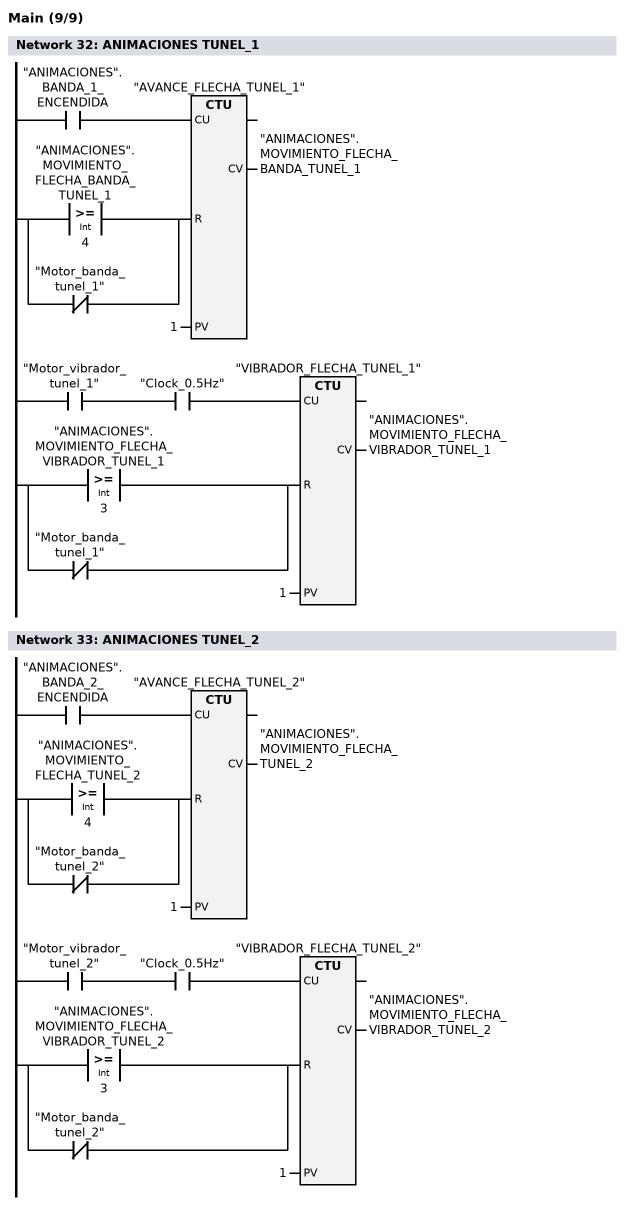
   "AVANCE_FLECHA_TUNEL_1".CTU(CU := "ANIMACIONES".BANDA_1_ENCENDIDA,
                           R := ("ANIMACIONES".MOVIMIENTO_FLECHA_BANDA_TUNEL_1 >= 4) OR NOT "Motor_banda_tunel_1",
                           PV := 1,
                           CV => "ANIMACIONES".MOVIMIENTO_FLECHA_BANDA_TUNEL_1);
   "VIBRADOR_FLECHA_TUNEL_1".CTU(CU := "Motor_vibrador_tunel_1" AND "Clock_0.5Hz",
                           R := ("ANIMACIONES".MOVIMIENTO_FLECHA_VIBRADOR_TUNEL_1 >= 3) OR NOT "Motor_banda_tunel_1",
                           PV := 1,
                           CV => "ANIMACIONES".MOVIMIENTO_FLECHA_VIBRADOR_TUNEL_1);
END_REGION

REGION Network 33: ANIMACIONES TUNEL_2
   "AVANCE_FLECHA_TUNEL_2".CTU(CU := "ANIMACIONES".BANDA_2_ENCENDIDA,
                           R := ("ANIMACIONES".MOVIMIENTO_FLECHA_TUNEL_2 >= 4) OR NOT "Motor_banda_tunel_2",
                           PV := 1,
                           CV => "ANIMACIONES".MOVIMIENTO_FLECHA_TUNEL_2);
   "VIBRADOR_FLECHA_TUNEL_2".CTU(CU := "Motor_vibrador_tunel_2" AND "Clock_0.5Hz",
                           R := ("ANIMACIONES".MOVIMIENTO_FLECHA_VIBRADOR_TUNEL_2 >= 3) OR NOT "Motor_banda_tunel_2",
                           PV := 1,
                           CV => "ANIMACIONES".MOVIMIENTO_FLECHA_VIBRADOR_TUNEL_2);
END_REGION
END_ORGANIZATION_BLOCK

(* ===== HMI "HMI_RT_1" =====
system functions are stored by id; their names below are inferred from use

HMI tags "Default tag table"
   "Tag_ScreenNumber" : UInt, internal

Template "Template_1" 800x480
   Button "Exit" at 714,429 size 71x50; TextOff 'Exit'; PictureOff "ExitRuntime_KTP700_Basic_PN_TR"; PictureOn "ExitRuntime_KTP700_Basic_PN_TR"
      on Release: StopRuntime(0)
   Button "Log on" at 614,429 size 71x50; TextOff 'Log on'; PictureOff "Login_KTP700_Basic_PN_TR"; PictureOn "Login_KTP700_Basic_PN_TR"
      on Release: function_a2a04561()
   Button "Template_Button" at 514,429 size 71x50; TextOff 'Text'
   Button "Template_Button_1" at 414,429 size 71x50; TextOff 'Text'
   Button "Template_Button_2" at 314,429 size 71x50; TextOff 'Text'
   Button "Template_Button_3" at 214,429 size 71x50; TextOff 'Text'
   Button "Alarms" at 114,429 size 71x50; TextOff 'Alarms'; PictureOff "AlarmDisplay_KTP700_Basic_PN_TR"; PictureOn "AlarmDisplay_KTP700_Basic_PN_TR"
      on Release: function_ef3f5d25("Alarm window_Unacknowledged", -1)
   Button "Start screen" at 14,429 size 71x50; TextOff 'Start screen'; PictureOff "NavigateHome_KTP700_Basic_PN_TR"; PictureOn "NavigateHome_KTP700_Basic_PN_TR"
      on Release: ActivateScreen("Root screen", 0)
   SymbolicIOField "Symbolic_IO_Field_Screen" at 93,9 size 600x33; TextOff '0'; TextOn '1'; TextList "TextList_ScreenNames"
      ProcessValue <- "Tag_ScreenNumber"
      on Change: ActivateScreenByNumber("Tag_ScreenNumber", 0)
   DateTimeField "HmiScreenItemData" at 695,25 size 105x25
   DateTimeField "HmiScreenItemData_1" at 695,0 size 105x25
   GraphicView "Logo" at 0,0 size 91x51; Picture "Logo of HMI_1"

screen "Root screen" 800x480, template "Template_1"
   on GenerateScreen: SetTag("Tag_ScreenNumber", 1)
   TextField "HmiScreenItemData" at 80,225 size 640x25; Text 'Welcome to HMI_1 (KTP700 Basic+ PN)!'
*)

(* ===== HMI "HMI_RT_2" =====
system functions are stored by id; their names below are inferred from use
connection "HMI_Connection_1": ETHERNET, SMART_S7_1500_OMS

HMI tags "Default tag table"
   "Tag_ScreenNumber" : UInt, internal
   "Motor_banda_tunel_1" : Bool = PLC Motor_banda_tunel_1 AT %Q10.0, 1 s
   "Señal_de_fallo_banda_tunel_1" : Bool = PLC Señal_de_fallo_banda_tunel_1 AT %I11.1, 1 s
   "PERMISOS_DE_MARCHA_TUNEL_1_BANDA_TUNEL_1_MANUAL" : Bool = PLC PERMISOS_DE_MARCHA_TUNEL_1.BANDA_TUNEL_1_MANUAL, 1 s
   "BOTONERA_HMI_TUNEL_1_KM1_INICIO_MANUAL_BANDA_TUNEL_1" : Bool = PLC BOTONERA_HMI_TUNEL_1.KM1_INICIO_MANUAL_BANDA_TUNEL_1, 1 s
   "BOTONERA_HMI_TUNEL_1_KM1_STOP_MANUAL_BANDA_TUNEL_1" : Bool = PLC BOTONERA_HMI_TUNEL_1.KM1_STOP_MANUAL_BANDA_TUNEL_1, 1 s
   "PERMISOS_DE_MARCHA_TUNEL_1_VENTILADOR_TUNEL_1_MANUAL" : Bool = PLC PERMISOS_DE_MARCHA_TUNEL_1.VENTILADOR_TUNEL_1_MANUAL, 1 s
   "Señal_de_fallo_ventilador_tunel_1" : Bool = PLC Señal_de_fallo_ventilador_tunel_1 AT %I11.3, 1 s
   "BOTONERA_HMI_TUNEL_1_KM2_INICIO_MANUAL_ASPIRADOR_TUNEL_1" : Bool = PLC BOTONERA_HMI_TUNEL_1.KM2_INICIO_MANUAL_ASPIRADOR_TUNEL_1, 1 s
   "BOTONERA_HMI_TUNEL_1_KM3_INICIO_MANUAL_VENTILADOR_TUNEL_1" : Bool = PLC BOTONERA_HMI_TUNEL_1.KM3_INICIO_MANUAL_VENTILADOR_TUNEL_1, 1 s
   "BOTONERA_HMI_TUNEL_1_KM3_STOP_MANUAL_VENTILADOR_TUNEL_1" : Bool = PLC BOTONERA_HMI_TUNEL_1.KM3_STOP_MANUAL_VENTILADOR_TUNEL_1, 1 s
   "PERMISOS_DE_MARCHA_TUNEL_1_ASPIRADOR_TUNEL_1_MANUAL" : Bool = PLC PERMISOS_DE_MARCHA_TUNEL_1.ASPIRADOR_TUNEL_1_MANUAL, 1 s
   "Señal_de_fallo_aspirador_tunel_1" : Bool = PLC Señal_de_fallo_aspirador_tunel_1 AT %I11.2, 1 s
   "BOTONERA_HMI_TUNEL_1_KM2_STOP_MANUAL_ASPIRADOR_TUNEL_1" : Bool = PLC BOTONERA_HMI_TUNEL_1.KM2_STOP_MANUAL_ASPIRADOR_TUNEL_1, 1 s
   "PERMISOS_DE_MARCHA_TUNEL_1_CERRAR_CUCHARA_TUNEL_1_MANUAL" : Bool = PLC PERMISOS_DE_MARCHA_TUNEL_1.CERRAR_CUCHARA_TUNEL_1_MANUAL, 1 s
   "PERMISOS_DE_MARCHA_TUNEL_1_ABRIR_CUCHARA_TUNEL_1_MANUAL" : Bool = PLC PERMISOS_DE_MARCHA_TUNEL_1.ABRIR_CUCHARA_TUNEL_1_MANUAL, 1 s
   "BOTONERA_HMI_TUNEL_1_SUBIR_CUCHARA_TUNEL_1" : Bool = PLC BOTONERA_HMI_TUNEL_1.SUBIR_CUCHARA_TUNEL_1, 1 s
   "BOTONERA_HMI_TUNEL_1_BAJAR_CUCHARA_TUNEL_1" : Bool = PLC BOTONERA_HMI_TUNEL_1.BAJAR_CUCHARA_TUNEL_1, 1 s
   "BOTONERA_HMI_TUNEL_1_CARGADOR_CAJAS_IZQUIERDA_TUNEL_1" : Bool = PLC BOTONERA_HMI_TUNEL_1.CARGADOR_CAJAS_IZQUIERDA_TUNEL_1, 1 s
   "PERMISOS_DE_MARCHA_TUNEL_1_CAJA_IZQUIERDA_TUNEL_1_MANUAL" : Bool = PLC PERMISOS_DE_MARCHA_TUNEL_1.CAJA_IZQUIERDA_TUNEL_1_MANUAL, 1 s
   "PERMISOS_DE_MARCHA_TUNEL_1_CAJA_DERECHA_TUNEL_1_MANUAL" : Bool = PLC PERMISOS_DE_MARCHA_TUNEL_1.CAJA_DERECHA_TUNEL_1_MANUAL, 1 s
   "BOTONERA_HMI_TUNEL_1_CARGADOR_CAJAS_DERECHA_TUNEL_1" : Bool = PLC BOTONERA_HMI_TUNEL_1.CARGADOR_CAJAS_DERECHA_TUNEL_1, 1 s
   "BOTONERA_HMI_TUNEL_1_KM4_INICIO_MANUAL_VIBRADOR_TUNEL_1" : Bool = PLC BOTONERA_HMI_TUNEL_1.KM4_INICIO_MANUAL_VIBRADOR_TUNEL_1, 1 s
   "BOTONERA_HMI_TUNEL_1_KM4_STOP_MANUAL_VIBRADOR_TUNEL_1" : Bool = PLC BOTONERA_HMI_TUNEL_1.KM4_STOP_MANUAL_VIBRADOR_TUNEL_1, 1 s
   "PERMISOS_DE_MARCHA_TUNEL_1_VIBRADOR_TUNEL_1_MANUAL" : Bool = PLC PERMISOS_DE_MARCHA_TUNEL_1.VIBRADOR_TUNEL_1_MANUAL, 1 s
   "Señal_de_fallo_vibrador_tunel_1" : Bool = PLC Señal_de_fallo_vibrador_tunel_1 AT %I11.4, 1 s
   "ANIMACIONES_MOVIMIENTO_FLECHA_TUNEL_1" : Int = PLC ANIMACIONES.MOVIMIENTO_FLECHA_BANDA_TUNEL_1, 1 s
   "ANIMACIONES_MOVIMIENTO_FLECHA_VIBRADOR_TUNEL_1" : Int = PLC ANIMACIONES.MOVIMIENTO_FLECHA_VIBRADOR_TUNEL_1, 1 s
   "Señalizacion_operacion_verde_tunel_1" : Bool = PLC Señalizacion_operacion_verde_tunel_1 AT %Q11.3, 1 s
   "Señalizacion_azul_tunel_1" : Bool = PLC Señalizacion_azul_tunel_1 AT %Q11.2, 1 s
   "Señalizacion_Roja_Tunel_1" : Bool = PLC Señalizacion_Roja_Tunel_1 AT %Q11.1, 1 s
   "PERMISOS_DE_MARCHA_TUNEL_1_VENTILADOR_TUNEL_1_AUTOMATICO" : Bool = PLC PERMISOS_DE_MARCHA_TUNEL_1.VENTILADOR_TUNEL_1_AUTOMATICO, 1 s
   "PERMISOS_DE_MARCHA_TUNEL_1_ASPIRADOR_TUNEL_1_AUTOMATICO" : Bool = PLC PERMISOS_DE_MARCHA_TUNEL_1.ASPIRADOR_TUNEL_1_AUTOMATICO, 1 s
   "PERMISOS_DE_MARCHA_TUNEL_1_BANDA_TUNEL_1_AUTOMATICO" : Bool = PLC PERMISOS_DE_MARCHA_TUNEL_1.BANDA_TUNEL_1_AUTOMATICO, 1 s
   "PERMISOS_DE_MARCHA_TUNEL_1_VIBRADOR_TUNEL_1_AUTOMATICO" : Bool = PLC PERMISOS_DE_MARCHA_TUNEL_1.VIBRADOR_TUNEL_1_AUTOMATICO, 1 s
   "PERMISOS_DE_MARCHA_TUNEL_1_CAJA_DERECHA_TUNEL_1_AUTOMATICO" : Bool = PLC PERMISOS_DE_MARCHA_TUNEL_1.CAJA_DERECHA_TUNEL_1_AUTOMATICO, 1 s
   "PERMISOS_DE_MARCHA_TUNEL_1_CAJA_IZQUIERDA_TUNEL_1_AUTOMATICO" : Bool = PLC PERMISOS_DE_MARCHA_TUNEL_1.CAJA_IZQUIERDA_TUNEL_1_AUTOMATICO, 1 s
   "PERMISOS_DE_MARCHA_TUNEL_1_CERRAR_CUCHARA_TUNEL_1_AUTOMATICO" : Bool = PLC PERMISOS_DE_MARCHA_TUNEL_1.CERRAR_CUCHARA_TUNEL_1_AUTOMATICO, 1 s
   "PERMISOS_DE_MARCHA_TUNEL_1_ABRIR_CUCHARA_TUNEL_1_AUTOMATICO" : Bool = PLC PERMISOS_DE_MARCHA_TUNEL_1.ABRIR_CUCHARA_TUNEL_1_AUTOMATICO, 1 s
   "Motor_aspirador_tunel_!" : Bool = PLC Motor_aspirador_tunel_! AT %Q10.1, 1 s
   "Motor_ventilador_tunel_1" : Bool = PLC Motor_ventilador_tunel_1 AT %Q10.2, 1 s
   "Motor_vibrador_tunel_1" : Bool = PLC Motor_vibrador_tunel_1 AT %Q10.3, 1 s
   "Subir_Cuchara_Tunel_1" : Bool = PLC Subir_Cuchara_Tunel_1 AT %Q11.0, 1 s
   "Bajar_cuchara_Tunel_1" : Bool = PLC Bajar_cuchara_Tunel_1 AT %Q10.7, 1 s
   "Desviar_cajas_derecha_Tunel_1" : Bool = PLC Desviar_cajas_derecha_Tunel_1 AT %Q10.4, 1 s
   "Desviar_cajas_izquierda_Tunel_1" : Bool = PLC Desviar_cajas_izquierda_Tunel_1 AT %Q10.5, 1 s
   "TEMPORIZADOR_PASO_TAPAS_TUNEL_1" : Int = PLC TEMPORIZADOR_PASO_TAPAS_TUNEL_1 AT %MW0, 1 s
   "TEMPORIZADOR_BLOQUEO_TAPAS_TUNEL_1" : Int = PLC TEMPORIZADOR_BLOQUEO_TAPAS_TUNEL_1 AT %MW2, 1 s
   "TEMPORIZADOR_CAMBIO_DE_LLENADO_CAJA_TUNEL_1" : Int = PLC TEMPORIZADOR_CAMBIO_DE_LLENADO_CAJA_TUNEL_1 AT %MW4, 1 s
   "PERMISOS_GENERALES_MODO_LOCAL_1" : Bool = PLC PERMISOS_GENERALES.MODO_LOCAL_1, 1 s
   "PERMISOS_GENERALES_MODO_AUTOMATICO_1" : Bool = PLC PERMISOS_GENERALES.MODO_AUTOMATICO_1, 1 s
   "ALARMAS_TUNEL_1" : Int AT %DB24.DBW0, 1 s

discrete alarms
   1: 'Revisar estado guardamotor QM1', class Errors, trigger "ALARMAS_TUNEL_1" bit 8
   2: 'Revisar estado guardamotor QM2', class Warnings, trigger "ALARMAS_TUNEL_1" bit 9
   3: 'Revisar estado guardamotor QM3', class Warnings, trigger "ALARMAS_TUNEL_1" bit 10
   4: 'Revisar estado guardamotor QM4', class Errors, trigger "ALARMAS_TUNEL_1" bit 11
   5: 'Revisar presion en red neumatica', class Errors, trigger "ALARMAS_TUNEL_1" bit 12
   6: 'Equipo en paro de emergencia', class Errors, trigger "ALARMAS_TUNEL_1" bit 14
   7: 'Sin suministro de tapas en entrada', class Warnings, trigger "ALARMAS_TUNEL_1" bit 13

Template "Template_1" 800x480
   Button "Exit" at 714,429 size 71x50; TextOff 'Exit'; PictureOff "ExitRuntime_KTP700_Basic_PN_TR"; PictureOn "ExitRuntime_KTP700_Basic_PN_TR"
      on Release: StopRuntime(0)
   Button "Log on" at 614,429 size 71x50; TextOff 'Log on'; PictureOff "Login_KTP700_Basic_PN_TR"; PictureOn "Login_KTP700_Basic_PN_TR"
      on Release: function_a2a04561()
   Button "Template_Button" at 514,429 size 71x50; TextOff 'Text'
   Button "Template_Button_1" at 414,429 size 71x50; TextOff 'Text'
   Button "Template_Button_2" at 314,429 size 71x50; TextOff 'Text'
   Button "Template_Button_3" at 214,429 size 71x50; TextOff 'Text'
   Button "Alarms" at 114,429 size 71x50; TextOff 'Alarms'; PictureOff "AlarmDisplay_KTP700_Basic_PN_TR"; PictureOn "AlarmDisplay_KTP700_Basic_PN_TR"
   Button "Start screen" at 14,429 size 71x50; TextOff 'Start screen'; PictureOff "NavigateHome_KTP700_Basic_PN_TR"; PictureOn "NavigateHome_KTP700_Basic_PN_TR"
      on Release: ActivateScreen("PANTALLA DE INICIO", 0)
   SymbolicIOField "Symbolic_IO_Field_Screen" at 93,9 size 600x33; TextOff '0'; TextOn '1'; TextList "TextList_ScreenNames"
      ProcessValue <- "Tag_ScreenNumber"
      on Change: ActivateScreenByNumber("Tag_ScreenNumber", 0)
   DateTimeField "HmiScreenItemData" at 695,25 size 105x25
   DateTimeField "HmiScreenItemData_1" at 695,0 size 105x25
   GraphicView "Logo" at 0,0 size 91x51; Picture "Logo of HMI_1"

screen "PANTALLA DE INICIO" 800x480, template "Template_1"
   on GenerateScreen: SetTag("Tag_ScreenNumber", 1)
   GraphicView "Graphic view_1" at 302,101 size 200x200; Picture "pngegg"
   Button "Button_1" at 277,47 size 251x30; TextOff 'TUNEL ENFRIAMIENTO 1'
   Button "Button_2" at 244,83 size 316x30; TextOff 'LINEA DE FABRICACION DE TAPAS 2'
   GraphicView "Graphic view_2" at 352,314 size 100x100; Picture "selector-de-llave-3-posiciones-enclavamiento-eaton-moeller-111774-m22-wrs3-ms3-removebg-preview"
   Button "Button_3" at 131,282 size 96x32; TextOff 'LOCAL'; Authorization "Mantenimiento"
      on Press: ActivateScreen("MODO LOCAL", 0)
   Button "Button_4" at 590,282 size 96x32; TextOff 'REMOTO'
      on Press: ActivateScreen("MODO REMOTO", 0)

screen "MODO LOCAL" 800x480
   GraphicView "Graphic view_8" at 402,218 size 50x50; Picture "Graphic_9"
      Visibility <- "PERMISOS_DE_MARCHA_TUNEL_1_VENTILADOR_TUNEL_1_MANUAL"
   GraphicView "Graphic view_1" at 0,0 size 100x100; Picture "pngegg"
   GraphicView "Graphic view_2" at 126,262 size 624x99; Picture "Graphic_1"
   GraphicView "Graphic view_3" at 470,311 size 50x50; Picture "Graphic_2"
      Visibility <- "PERMISOS_DE_MARCHA_TUNEL_1_BANDA_TUNEL_1_MANUAL"
   GraphicView "Graphic view_4" at 470,311 size 50x50; Picture "Graphic_3"
      Visibility <- "Motor_banda_tunel_1"
   GraphicView "Graphic view_5" at 470,311 size 50x50; Picture "Graphic_4"
      Visibility <- "Señal_de_fallo_banda_tunel_1"
   Button "Button_2" at 466,363 size 50x20; TextOff 'ON'; Authorization "Mantenimiento"
      on Press: SetBit("BOTONERA_HMI_TUNEL_1_KM1_INICIO_MANUAL_BANDA_TUNEL_1")
      on Release: ResetBit("BOTONERA_HMI_TUNEL_1_KM1_INICIO_MANUAL_BANDA_TUNEL_1")
      Visibility <- "PERMISOS_GENERALES_MODO_LOCAL_1"
   Button "Button_3" at 522,362 size 50x20; TextOff 'OFF'; Authorization "Mantenimiento"
      on Press: SetBit("BOTONERA_HMI_TUNEL_1_KM1_STOP_MANUAL_BANDA_TUNEL_1")
      on Release: ResetBit("BOTONERA_HMI_TUNEL_1_KM1_STOP_MANUAL_BANDA_TUNEL_1")
      Visibility <- "PERMISOS_GENERALES_MODO_LOCAL_1"
   GraphicView "Graphic view_6" at 401,217 size 50x50; Picture "Graphic_6"
      Visibility <- "PERMISOS_DE_MARCHA_TUNEL_1_VENTILADOR_TUNEL_1_MANUAL"
   GraphicView "Graphic view_9" at 356,222 size 48x45; Picture "viento"
      Visibility <- "PERMISOS_DE_MARCHA_TUNEL_1_VENTILADOR_TUNEL_1_MANUAL"
   GraphicView "Graphic view_7" at 401,218 size 50x50; Picture "Graphic_7"
      Visibility <- "Señal_de_fallo_ventilador_tunel_1"
   Button "Button_1" at 359,194 size 50x20; TextOff 'ON'; Authorization "Mantenimiento"
      on Release: ResetBit("BOTONERA_HMI_TUNEL_1_KM3_INICIO_MANUAL_VENTILADOR_TUNEL_1")
      on Press: SetBit("BOTONERA_HMI_TUNEL_1_KM3_INICIO_MANUAL_VENTILADOR_TUNEL_1")
   Button "Button_4" at 419,195 size 50x20; TextOff 'OFF'; Authorization "Mantenimiento"
      on Release: ResetBit("BOTONERA_HMI_TUNEL_1_KM3_STOP_MANUAL_VENTILADOR_TUNEL_1")
      on Press: SetBit("BOTONERA_HMI_TUNEL_1_KM3_STOP_MANUAL_VENTILADOR_TUNEL_1")
   GraphicView "Graphic view_10" at 240,300 size 50x50; Picture "Graphic_23"
      Visibility <- "PERMISOS_DE_MARCHA_TUNEL_1_ASPIRADOR_TUNEL_1_MANUAL"
   GraphicView "Graphic view_11" at 240,300 size 50x50; Picture "Graphic_24"
      Visibility <- "PERMISOS_DE_MARCHA_TUNEL_1_ASPIRADOR_TUNEL_1_MANUAL"
   GraphicView "Graphic view_12" at 240,300 size 50x50; Picture "Graphic_25"
      Visibility <- "Señal_de_fallo_aspirador_tunel_1"
   GraphicView "Graphic view_13" at 209,321 size 52x87; Picture "viento"
      Visibility <- "PERMISOS_DE_MARCHA_TUNEL_1_ASPIRADOR_TUNEL_1_MANUAL"
   Button "Button_5" at 211,388 size 50x20; TextOff 'ON'; Authorization "Mantenimiento"
      on Release: ResetBit("BOTONERA_HMI_TUNEL_1_KM2_INICIO_MANUAL_ASPIRADOR_TUNEL_1")
      on Press: SetBit("BOTONERA_HMI_TUNEL_1_KM2_INICIO_MANUAL_ASPIRADOR_TUNEL_1")
   Button "Button_6" at 265,389 size 50x20; TextOff 'OFF'; Authorization "Mantenimiento"
      on Release: ResetBit("BOTONERA_HMI_TUNEL_1_KM2_STOP_MANUAL_ASPIRADOR_TUNEL_1")
      on Press: SetBit("BOTONERA_HMI_TUNEL_1_KM2_STOP_MANUAL_ASPIRADOR_TUNEL_1")
   TextField "Text field_1" at 463,386 size 109x23; Text 'Motor Banda'
   TextField "Text field_2" at 376,159 size 90x23; Text 'Ventilador'
   TextField "Text field_3" at 231,411 size 81x23; Text 'Extractor'
   GraphicView "Graphic view_15" at 500,76 size 300x200; Picture "Compuerta"
      Visibility <- "PERMISOS_DE_MARCHA_TUNEL_1_ABRIR_CUCHARA_TUNEL_1_MANUAL"
   GraphicView "Graphic view_14" at 499,139 size 300x200; Picture "Compuerta"
      Visibility <- "PERMISOS_DE_MARCHA_TUNEL_1_CERRAR_CUCHARA_TUNEL_1_MANUAL"
   Button "Button_7" at 724,120 size 60x20; TextOff 'SUBIR'; Authorization "Mantenimiento"
      on Release: ResetBit("BOTONERA_HMI_TUNEL_1_SUBIR_CUCHARA_TUNEL_1")
      on Press: SetBit("BOTONERA_HMI_TUNEL_1_SUBIR_CUCHARA_TUNEL_1")
      Appearance <- "PERMISOS_DE_MARCHA_TUNEL_1_ABRIR_CUCHARA_TUNEL_1_MANUAL"
   Button "Button_8" at 724,154 size 60x20; TextOff 'BAJAR'; Authorization "Mantenimiento"
      on Release: ResetBit("BOTONERA_HMI_TUNEL_1_BAJAR_CUCHARA_TUNEL_1")
      on Press: SetBit("BOTONERA_HMI_TUNEL_1_BAJAR_CUCHARA_TUNEL_1")
      Appearance <- "PERMISOS_DE_MARCHA_TUNEL_1_CERRAR_CUCHARA_TUNEL_1_MANUAL"
   Button "Button_9" at 16,155 size 100x20; TextOff 'IZQUIERDA'; Authorization "Mantenimiento"
      on Release: ResetBit("BOTONERA_HMI_TUNEL_1_CARGADOR_CAJAS_IZQUIERDA_TUNEL_1")
      on Press: SetBit("BOTONERA_HMI_TUNEL_1_CARGADOR_CAJAS_IZQUIERDA_TUNEL_1")
      Appearance <- "PERMISOS_DE_MARCHA_TUNEL_1_CAJA_IZQUIERDA_TUNEL_1_MANUAL"
   Button "Button_10" at 169,155 size 100x20; TextOff 'DERECHA'; Authorization "Mantenimiento"
      on Release: ResetBit("BOTONERA_HMI_TUNEL_1_CARGADOR_CAJAS_DERECHA_TUNEL_1")
      on Press: SetBit("BOTONERA_HMI_TUNEL_1_CARGADOR_CAJAS_DERECHA_TUNEL_1")
      Appearance <- "PERMISOS_DE_MARCHA_TUNEL_1_CAJA_DERECHA_TUNEL_1_MANUAL"
   Button "Button_11" at 400,440 size 368x32; TextOff 'ESTADO DE ELEMENTOS Y ACTUADORES'
      on Press: ActivateScreen("VISUALIZACION DE ESTADOS LOCAL TUNEL 1", 0)
   TextField "Text field_4" at 229,86 size 241x33; Text 'MODO LOCAL ACTIVO'
   GraphicView "Graphic view_16" at 496,268 size 87x56; Picture "pngtree-vector-back-icon-png-image_956547-removebg-preview"
      Visibility <- "ANIMACIONES_MOVIMIENTO_FLECHA_TUNEL_1"
   GraphicView "Graphic view_17" at 210,262 size 87x56; Picture "pngtree-vector-back-icon-png-image_956547-removebg-preview"
      Visibility <- "ANIMACIONES_MOVIMIENTO_FLECHA_TUNEL_1"
   GraphicView "Graphic view_18" at 350,266 size 87x56; Picture "pngtree-vector-back-icon-png-image_956547-removebg-preview"
      Visibility <- "ANIMACIONES_MOVIMIENTO_FLECHA_TUNEL_1"
   GraphicView "Graphic view_19" at 0,296 size 209x184; Picture "AGITADOR"
   GraphicView "Graphic view_20" at 16,418 size 50x50; Picture "Graphic_4"
      Visibility <- "Señal_de_fallo_vibrador_tunel_1"
   GraphicView "Graphic view_21" at 16,417 size 50x50; Picture "Graphic_2"
      Visibility <- "PERMISOS_DE_MARCHA_TUNEL_1_VIBRADOR_TUNEL_1_MANUAL"
   GraphicView "Graphic view_22" at 16,416 size 50x50; Picture "Graphic_3"
      Visibility <- "PERMISOS_DE_MARCHA_TUNEL_1_VIBRADOR_TUNEL_1_MANUAL"
   GraphicView "Graphic view_23" at 4,366 size 35x40; Picture "FLECHA ARRIBA"
      Visibility <- "ANIMACIONES_MOVIMIENTO_FLECHA_VIBRADOR_TUNEL_1"
   GraphicView "Graphic view_24" at 160,366 size 35x40; Picture "FLECHA ABAJO"
      Visibility <- "ANIMACIONES_MOVIMIENTO_FLECHA_VIBRADOR_TUNEL_1"
   GraphicView "Graphic view_25" at 160,366 size 35x40; Picture "FLECHA ARRIBA"
      Visibility <- "ANIMACIONES_MOVIMIENTO_FLECHA_VIBRADOR_TUNEL_1"
   GraphicView "Graphic view_26" at 4,366 size 35x40; Picture "FLECHA ABAJO"
      Visibility <- "ANIMACIONES_MOVIMIENTO_FLECHA_VIBRADOR_TUNEL_1"
   GraphicView "Graphic view_27" at 0,192 size 119x73; Picture "CAJA_1"
      Visibility <- "PERMISOS_DE_MARCHA_TUNEL_1_CAJA_IZQUIERDA_TUNEL_1_MANUAL"
   GraphicView "Graphic view_28" at 160,192 size 119x73; Picture "CAJA_1"
      Visibility <- "PERMISOS_DE_MARCHA_TUNEL_1_CAJA_DERECHA_TUNEL_1_MANUAL"
   GraphicView "Graphic view_29" at 712,14 size 60x60; Picture "Graphic_28"
      Visibility <- "Señalizacion_operacion_verde_tunel_1"
   GraphicView "Graphic view_30" at 714,14 size 60x60; Picture "Graphic_29"
      Visibility <- "Señalizacion_azul_tunel_1"
   GraphicView "Graphic view_31" at 716,14 size 60x60; Picture "Graphic_31"
      Visibility <- "Señalizacion_Roja_Tunel_1"
   Button "Button_12" at 14,320 size 50x20; TextOff 'ON'; Authorization "Mantenimiento"
      on Release: ResetBit("BOTONERA_HMI_TUNEL_1_KM4_INICIO_MANUAL_VIBRADOR_TUNEL_1")
      on Press: SetBit("BOTONERA_HMI_TUNEL_1_KM4_INICIO_MANUAL_VIBRADOR_TUNEL_1")
   Button "Button_13" at 75,319 size 50x20; TextOff 'OFF'; Authorization "Mantenimiento"
      on Release: ResetBit("BOTONERA_HMI_TUNEL_1_KM4_STOP_MANUAL_VIBRADOR_TUNEL_1")
      on Press: SetBit("BOTONERA_HMI_TUNEL_1_KM4_STOP_MANUAL_VIBRADOR_TUNEL_1")
   TextField "Text field_5" at 35,292 size 75x23; Text 'Vibrador'
   UserView "User view_1" at 118,10 size 564x55
   Softkey "Softkey_F1" at 0,0 size 0x0
      on KeyDown: ActivateScreen("PANTALLA DE INICIO", 0)

screen "VISUALIZACION DE ESTADOS LOCAL TUNEL 1" 800x480
   GraphicView "Graphic view_1" at 0,0 size 100x100; Picture "pngegg"
   Button "Button_11" at 223,435 size 368x32; TextOff 'VISUALIZACION MIMICO'
      on Press: ActivateScreen("MODO LOCAL", 0)
   TextField "Text field_4" at 259,75 size 322x43; Text 'MODO LOCAL ACTIVO'
   Button "Button_1" at 43,120 size 261x32; TextOff 'BANDA TRANSPORTADORA'
   Button "Button_2" at 43,169 size 261x32; TextOff 'EXTRACTOR'
   Button "Button_3" at 43,218 size 261x32; TextOff 'VENTILADOR'
   Button "Button_4" at 43,263 size 261x32; TextOff 'VIBRADOR'
   Button "Button_5" at 43,308 size 261x32; TextOff 'CUCHARA'
   Button "Button_6" at 43,353 size 261x32; TextOff 'CAJA'
   Button "Button_7" at 345,120 size 96x32; TextOff 'ON'; Authorization "Mantenimiento"
      on Press: SetBit("BOTONERA_HMI_TUNEL_1_KM1_INICIO_MANUAL_BANDA_TUNEL_1")
      on Release: ResetBit("BOTONERA_HMI_TUNEL_1_KM1_INICIO_MANUAL_BANDA_TUNEL_1")
   Button "Button_8" at 469,121 size 96x32; TextOff 'OFF'; Authorization "Mantenimiento"
      on Press: SetBit("BOTONERA_HMI_TUNEL_1_KM1_STOP_MANUAL_BANDA_TUNEL_1")
      on Release: ResetBit("BOTONERA_HMI_TUNEL_1_KM1_STOP_MANUAL_BANDA_TUNEL_1")
   Button "Button_9" at 604,121 size 96x32; TextOff 'APAGADO'
      Visibility <- "PERMISOS_DE_MARCHA_TUNEL_1_BANDA_TUNEL_1_MANUAL"
   Button "Button_10" at 601,120 size 106x32; TextOff 'ENCENDIDO'
      Visibility <- "PERMISOS_DE_MARCHA_TUNEL_1_BANDA_TUNEL_1_MANUAL"
   Button "Button_12" at 345,169 size 96x32; TextOff 'ON'; Authorization "Mantenimiento"
      on Release: ResetBit("BOTONERA_HMI_TUNEL_1_KM2_INICIO_MANUAL_ASPIRADOR_TUNEL_1")
      on Press: SetBit("BOTONERA_HMI_TUNEL_1_KM2_INICIO_MANUAL_ASPIRADOR_TUNEL_1")
   Button "Button_13" at 469,170 size 96x32; TextOff 'OFF'; Authorization "Mantenimiento"
      on Release: ResetBit("BOTONERA_HMI_TUNEL_1_KM2_STOP_MANUAL_ASPIRADOR_TUNEL_1")
      on Press: SetBit("BOTONERA_HMI_TUNEL_1_KM2_STOP_MANUAL_ASPIRADOR_TUNEL_1")
   Button "Button_14" at 604,170 size 96x32; TextOff 'APAGADO'
      Visibility <- "PERMISOS_DE_MARCHA_TUNEL_1_ASPIRADOR_TUNEL_1_MANUAL"
   Button "Button_15" at 601,169 size 106x32; TextOff 'ENCENDIDO'
      Visibility <- "PERMISOS_DE_MARCHA_TUNEL_1_ASPIRADOR_TUNEL_1_MANUAL"
   Button "Button_16" at 345,218 size 96x32; TextOff 'ON'; Authorization "Mantenimiento"
      on Release: ResetBit("BOTONERA_HMI_TUNEL_1_KM3_INICIO_MANUAL_VENTILADOR_TUNEL_1")
      on Press: SetBit("BOTONERA_HMI_TUNEL_1_KM3_STOP_MANUAL_VENTILADOR_TUNEL_1")
   Button "Button_17" at 469,219 size 96x32; TextOff 'OFF'; Authorization "Mantenimiento"
      on Release: ResetBit("BOTONERA_HMI_TUNEL_1_KM3_STOP_MANUAL_VENTILADOR_TUNEL_1")
      on Press: SetBit("BOTONERA_HMI_TUNEL_1_KM3_STOP_MANUAL_VENTILADOR_TUNEL_1")
   Button "Button_18" at 604,219 size 96x32; TextOff 'APAGADO'
      Visibility <- "PERMISOS_DE_MARCHA_TUNEL_1_VENTILADOR_TUNEL_1_MANUAL"
   Button "Button_19" at 601,219 size 106x32; TextOff 'ENCENDIDO'
      Visibility <- "PERMISOS_DE_MARCHA_TUNEL_1_VENTILADOR_TUNEL_1_MANUAL"
   Button "Button_20" at 345,267 size 96x32; TextOff 'ON'; Authorization "Mantenimiento"
      on Release: ResetBit("BOTONERA_HMI_TUNEL_1_KM4_INICIO_MANUAL_VIBRADOR_TUNEL_1")
      on Press: SetBit("BOTONERA_HMI_TUNEL_1_KM4_INICIO_MANUAL_VIBRADOR_TUNEL_1")
   Button "Button_21" at 469,268 size 96x32; TextOff 'OFF'; Authorization "Mantenimiento"
      on Release: ResetBit("BOTONERA_HMI_TUNEL_1_KM4_STOP_MANUAL_VIBRADOR_TUNEL_1")
      on Press: SetBit("BOTONERA_HMI_TUNEL_1_KM4_STOP_MANUAL_VIBRADOR_TUNEL_1")
   Button "Button_22" at 604,268 size 96x32; TextOff 'APAGADO'
      Visibility <- "PERMISOS_DE_MARCHA_TUNEL_1_VIBRADOR_TUNEL_1_MANUAL"
   Button "Button_23" at 601,267 size 106x32; TextOff 'ENCENDIDO'
      Visibility <- "PERMISOS_DE_MARCHA_TUNEL_1_VIBRADOR_TUNEL_1_MANUAL"
   Button "Button_24" at 345,308 size 96x32; TextOff 'ABRIR'; Authorization "Mantenimiento"
      on Release: ResetBit("BOTONERA_HMI_TUNEL_1_KM4_INICIO_MANUAL_VIBRADOR_TUNEL_1")
      on Press: SetBit("BOTONERA_HMI_TUNEL_1_KM4_INICIO_MANUAL_VIBRADOR_TUNEL_1")
   Button "Button_25" at 469,309 size 96x32; TextOff 'CERRAR'; Authorization "Mantenimiento"
      on Release: ResetBit("BOTONERA_HMI_TUNEL_1_KM4_STOP_MANUAL_VIBRADOR_TUNEL_1")
      on Press: SetBit("BOTONERA_HMI_TUNEL_1_KM4_STOP_MANUAL_VIBRADOR_TUNEL_1")
   Button "Button_26" at 604,309 size 96x32; TextOff 'ABIERTO'
      Visibility <- "PERMISOS_DE_MARCHA_TUNEL_1_ABRIR_CUCHARA_TUNEL_1_MANUAL"
   Button "Button_27" at 604,308 size 96x32; TextOff 'CERRADA'
      Visibility <- "PERMISOS_DE_MARCHA_TUNEL_1_CERRAR_CUCHARA_TUNEL_1_MANUAL"
   Button "Button_28" at 345,352 size 96x32; TextOff 'DERECHA'; Authorization "Mantenimiento"
      on Release: ResetBit("BOTONERA_HMI_TUNEL_1_KM4_INICIO_MANUAL_VIBRADOR_TUNEL_1")
      on Press: SetBit("BOTONERA_HMI_TUNEL_1_KM4_INICIO_MANUAL_VIBRADOR_TUNEL_1")
   Button "Button_29" at 469,353 size 96x32; TextOff 'IZQUIERDA'; Authorization "Mantenimiento"
      on Release: ResetBit("BOTONERA_HMI_TUNEL_1_KM4_STOP_MANUAL_VIBRADOR_TUNEL_1")
      on Press: SetBit("BOTONERA_HMI_TUNEL_1_KM4_STOP_MANUAL_VIBRADOR_TUNEL_1")
   Button "Button_30" at 604,353 size 96x32; TextOff 'DERECHA'
      Visibility <- "PERMISOS_DE_MARCHA_TUNEL_1_CAJA_DERECHA_TUNEL_1_MANUAL"
   Button "Button_31" at 601,351 size 96x32; TextOff 'IZQUIERDA'
      Visibility <- "PERMISOS_DE_MARCHA_TUNEL_1_CAJA_IZQUIERDA_TUNEL_1_MANUAL"
   GraphicView "Graphic view_2" at 729,118 size 35x35; Picture "ADVERTENCIA"
      Visibility <- "Señal_de_fallo_banda_tunel_1"
   GraphicView "Graphic view_3" at 729,166 size 35x35; Picture "ADVERTENCIA"
      Visibility <- "Señal_de_fallo_aspirador_tunel_1"
   GraphicView "Graphic view_4" at 729,214 size 35x35; Picture "ADVERTENCIA"
      Visibility <- "Señal_de_fallo_ventilador_tunel_1"
   GraphicView "Graphic view_5" at 729,264 size 35x35; Picture "ADVERTENCIA"
      Visibility <- "Señal_de_fallo_vibrador_tunel_1"
   UserView "User view_1" at 118,10 size 564x55
   Softkey "Softkey_F1" at 0,0 size 0x0
      on KeyDown: ActivateScreen("PANTALLA DE INICIO", 0)

screen "MODO REMOTO" 800x480
   TextField "Text field_4" at 229,86 size 267x33; Text 'MODO REMOTO ACTIVO'
   GraphicView "Graphic view_19" at 0,296 size 209x184; Picture "AGITADOR"
   GraphicView "Graphic view_2" at 126,262 size 624x99; Picture "Graphic_1"
   GraphicView "Graphic view_3" at 470,311 size 50x50; Picture "Graphic_2"
      Visibility <- "PERMISOS_DE_MARCHA_TUNEL_1_BANDA_TUNEL_1_AUTOMATICO"
   GraphicView "Graphic view_4" at 470,311 size 50x50; Picture "Graphic_3"
      Visibility <- "PERMISOS_DE_MARCHA_TUNEL_1_BANDA_TUNEL_1_AUTOMATICO"
   GraphicView "Graphic view_5" at 470,311 size 50x50; Picture "Graphic_4"
      Visibility <- "Señal_de_fallo_banda_tunel_1"
   GraphicView "Graphic view_6" at 401,217 size 50x50; Picture "Graphic_6"
      Visibility <- "PERMISOS_DE_MARCHA_TUNEL_1_VENTILADOR_TUNEL_1_AUTOMATICO"
   GraphicView "Graphic view_9" at 356,222 size 48x45; Picture "viento"
      Visibility <- "PERMISOS_DE_MARCHA_TUNEL_1_VENTILADOR_TUNEL_1_AUTOMATICO"
   GraphicView "Graphic view_8" at 401,218 size 50x50; Picture "Graphic_9"
      Visibility <- "PERMISOS_DE_MARCHA_TUNEL_1_VENTILADOR_TUNEL_1_AUTOMATICO"
   GraphicView "Graphic view_10" at 240,300 size 50x50; Picture "Graphic_23"
      Visibility <- "PERMISOS_DE_MARCHA_TUNEL_1_ASPIRADOR_TUNEL_1_AUTOMATICO"
   GraphicView "Graphic view_11" at 240,300 size 50x50; Picture "Graphic_24"
      Visibility <- "PERMISOS_DE_MARCHA_TUNEL_1_ASPIRADOR_TUNEL_1_AUTOMATICO"
   GraphicView "Graphic view_12" at 240,300 size 50x50; Picture "Graphic_25"
      Visibility <- "Señal_de_fallo_aspirador_tunel_1"
   GraphicView "Graphic view_13" at 211,335 size 52x55; Picture "viento"
      Visibility <- "PERMISOS_DE_MARCHA_TUNEL_1_BANDA_TUNEL_1_AUTOMATICO"
   TextField "Text field_1" at 444,363 size 109x23; Text 'Motor Banda'
   TextField "Text field_2" at 374,194 size 90x23; Text 'Ventilador'
   TextField "Text field_3" at 261,350 size 81x23; Text 'Extractor'
   Button "Button_7" at 718,120 size 78x20; TextOff 'ABIERTO'
      on Release: ResetBit("BOTONERA_HMI_TUNEL_1_SUBIR_CUCHARA_TUNEL_1")
      on Press: SetBit("BOTONERA_HMI_TUNEL_1_SUBIR_CUCHARA_TUNEL_1")
      Visibility <- "PERMISOS_DE_MARCHA_TUNEL_1_ABRIR_CUCHARA_TUNEL_1_AUTOMATICO"
   Button "Button_8" at 716,120 size 81x20; TextOff 'CERRADO'
      on Release: ResetBit("BOTONERA_HMI_TUNEL_1_BAJAR_CUCHARA_TUNEL_1")
      on Press: SetBit("BOTONERA_HMI_TUNEL_1_BAJAR_CUCHARA_TUNEL_1")
      Visibility <- "PERMISOS_DE_MARCHA_TUNEL_1_CERRAR_CUCHARA_TUNEL_1_AUTOMATICO"
   Button "Button_9" at 16,155 size 100x20; TextOff 'IZQUIERDA'
      Visibility <- "PERMISOS_DE_MARCHA_TUNEL_1_CAJA_IZQUIERDA_TUNEL_1_AUTOMATICO"
   Button "Button_10" at 169,155 size 100x20; TextOff 'DERECHA'
      Visibility <- "PERMISOS_DE_MARCHA_TUNEL_1_CAJA_DERECHA_TUNEL_1_AUTOMATICO"
   Button "Button_11" at 400,440 size 368x32; TextOff 'ESTADO DE ELEMENTOS Y ACTUADORES'
      on Press: ActivateScreen("VISUALIZACION DE ESTADOS LOCAL TUNEL 1", 0)
   GraphicView "Graphic view_16" at 496,268 size 87x56; Picture "pngtree-vector-back-icon-png-image_956547-removebg-preview"
      Visibility <- "ANIMACIONES_MOVIMIENTO_FLECHA_TUNEL_1"
   GraphicView "Graphic view_17" at 210,262 size 87x56; Picture "pngtree-vector-back-icon-png-image_956547-removebg-preview"
      Visibility <- "ANIMACIONES_MOVIMIENTO_FLECHA_TUNEL_1"
   GraphicView "Graphic view_18" at 350,266 size 87x56; Picture "pngtree-vector-back-icon-png-image_956547-removebg-preview"
      Visibility <- "ANIMACIONES_MOVIMIENTO_FLECHA_TUNEL_1"
   GraphicView "Graphic view_21" at 16,418 size 50x50; Picture "Graphic_2"
      Visibility <- "PERMISOS_DE_MARCHA_TUNEL_1_VIBRADOR_TUNEL_1_AUTOMATICO"
   GraphicView "Graphic view_22" at 17,417 size 50x50; Picture "Graphic_3"
      Visibility <- "PERMISOS_DE_MARCHA_TUNEL_1_VIBRADOR_TUNEL_1_AUTOMATICO"
   GraphicView "Graphic view_23" at 4,366 size 35x40; Picture "FLECHA ARRIBA"
      Visibility <- "ANIMACIONES_MOVIMIENTO_FLECHA_VIBRADOR_TUNEL_1"
   GraphicView "Graphic view_24" at 160,366 size 35x40; Picture "FLECHA ABAJO"
      Visibility <- "ANIMACIONES_MOVIMIENTO_FLECHA_VIBRADOR_TUNEL_1"
   GraphicView "Graphic view_25" at 160,366 size 35x40; Picture "FLECHA ARRIBA"
      Visibility <- "ANIMACIONES_MOVIMIENTO_FLECHA_VIBRADOR_TUNEL_1"
   GraphicView "Graphic view_26" at 4,366 size 35x40; Picture "FLECHA ABAJO"
      Visibility <- "ANIMACIONES_MOVIMIENTO_FLECHA_VIBRADOR_TUNEL_1"
   GraphicView "Graphic view_27" at 0,192 size 119x73; Picture "CAJA_1"
      Visibility <- "PERMISOS_DE_MARCHA_TUNEL_1_CAJA_IZQUIERDA_TUNEL_1_AUTOMATICO"
   GraphicView "Graphic view_28" at 160,192 size 119x73; Picture "CAJA_1"
      Visibility <- "PERMISOS_DE_MARCHA_TUNEL_1_CAJA_DERECHA_TUNEL_1_AUTOMATICO"
   GraphicView "Graphic view_29" at 712,14 size 60x60; Picture "Graphic_28"
      Visibility <- "Señalizacion_operacion_verde_tunel_1"
   GraphicView "Graphic view_30" at 714,14 size 60x60; Picture "Graphic_29"
      Visibility <- "Señalizacion_azul_tunel_1"
   GraphicView "Graphic view_31" at 716,14 size 60x60; Picture "Graphic_31"
      Visibility <- "Señalizacion_Roja_Tunel_1"
   TextField "Text field_5" at 33,310 size 75x23; Text 'Vibrador'
   GraphicView "Graphic view_7" at 401,218 size 50x50; Picture "Graphic_7"
      Visibility <- "Señal_de_fallo_ventilador_tunel_1"
   GraphicView "Graphic view_20" at 16,418 size 50x50; Picture "Graphic_4"
      Visibility <- "Señal_de_fallo_vibrador_tunel_1"
   GraphicView "Graphic view_14" at 500,125 size 300x200; Picture "Compuerta"
      Visibility <- "PERMISOS_DE_MARCHA_TUNEL_1_CERRAR_CUCHARA_TUNEL_1_AUTOMATICO"
   GraphicView "Graphic view_15" at 500,73 size 300x200; Picture "Compuerta"
      Visibility <- "PERMISOS_DE_MARCHA_TUNEL_1_ABRIR_CUCHARA_TUNEL_1_AUTOMATICO"
   Button "Button_5" at 279,376 size 50x20; TextOff 'ON'
      Visibility <- "Motor_aspirador_tunel_!"
   Button "Button_4" at 279,375 size 50x20; TextOff 'OFF'
      Visibility <- "Motor_aspirador_tunel_!"
   Button "Button_1" at 470,390 size 50x20; TextOff 'OFF'
      Visibility <- "Motor_banda_tunel_1"
   Button "Button_2" at 470,389 size 50x20; TextOff 'ON'
      Visibility <- "Motor_banda_tunel_1"
   GraphicView "Graphic view_1" at 341,344 size 41x39; Picture "ADVERTENCIA"
      Visibility <- "Señal_de_fallo_aspirador_tunel_1"
   GraphicView "Graphic view_32" at 549,352 size 41x39; Picture "ADVERTENCIA"
      Visibility <- "Señal_de_fallo_banda_tunel_1"
   Button "Button_3" at 392,172 size 50x20; TextOff 'ON'
      Visibility <- "Motor_ventilador_tunel_1"
   Button "Button_6" at 393,172 size 50x20; TextOff 'OFF'
      Visibility <- "Motor_ventilador_tunel_1"
   GraphicView "Graphic view_33" at 458,185 size 41x39; Picture "ADVERTENCIA"
      Visibility <- "Señal_de_fallo_ventilador_tunel_1"
   Button "Button_12" at 45,286 size 50x20; TextOff 'OFF'
      Visibility <- "Motor_vibrador_tunel_1"
   Button "Button_13" at 44,286 size 50x20; TextOff 'ON'
      Visibility <- "Motor_vibrador_tunel_1"
   GraphicView "Graphic view_34" at 106,295 size 41x39; Picture "ADVERTENCIA"
      Visibility <- "Señal_de_fallo_vibrador_tunel_1"
   GraphicView "Graphic view_35" at 0,0 size 100x100; Picture "pngegg"
   Button "Button_14" at 209,439 size 172x32; TextOff 'CONFIGURACION'; Authorization "Mantenimiento"
      on Press: ActivateScreen("VISUALIZACION DE ESTADOS LOCAL TUNEL 1", 0)
   UserView "User view_1" at 118,10 size 564x55
   Softkey "Softkey_F1" at 0,0 size 0x0
      on KeyDown: ActivateScreen("PANTALLA DE INICIO", 0)

screen "VISUALIZACION DE ESTADOS REMOTO TUNEL 1" 800x480
   Button "Button_1" at 43,120 size 261x32; TextOff 'BANDA TRANSPORTADORA'
   Button "Button_2" at 43,169 size 261x32; TextOff 'EXTRACTOR'
   Button "Button_3" at 43,218 size 261x32; TextOff 'VENTILADOR'
   Button "Button_4" at 43,263 size 261x32; TextOff 'VIBRADOR'
   Button "Button_5" at 43,308 size 261x32; TextOff 'CUCHARA'
   Button "Button_6" at 43,353 size 261x32; TextOff 'CAJA'
   Button "Button_7" at 345,120 size 96x32; TextOff 'ON'
      Visibility <- "Motor_banda_tunel_1"
   Button "Button_8" at 469,121 size 96x32; TextOff 'OFF'
      on Release: ResetBit("BOTONERA_HMI_TUNEL_1_KM1_STOP_MANUAL_BANDA_TUNEL_1")
      on Press: SetBit("BOTONERA_HMI_TUNEL_1_KM1_STOP_MANUAL_BANDA_TUNEL_1")
      Visibility <- "Motor_banda_tunel_1"
   Button "Button_9" at 604,121 size 96x32; TextOff 'FALLA'
      Visibility <- "Señal_de_fallo_banda_tunel_1"
   Button "Button_12" at 345,169 size 96x32; TextOff 'ON'
      Visibility <- "Motor_aspirador_tunel_!"
   Button "Button_13" at 469,170 size 96x32; TextOff 'OFF'
      Visibility <- "Motor_aspirador_tunel_!"
   Button "Button_14" at 604,170 size 96x32; TextOff 'FALLA'
      Visibility <- "Señal_de_fallo_aspirador_tunel_1"
   Button "Button_16" at 345,218 size 96x32; TextOff 'ON'
      Visibility <- "Motor_ventilador_tunel_1"
   Button "Button_17" at 469,219 size 96x32; TextOff 'OFF'
      Visibility <- "Motor_ventilador_tunel_1"
   Button "Button_18" at 604,219 size 96x32; TextOff 'FALLA'
      Visibility <- "Señal_de_fallo_ventilador_tunel_1"
   Button "Button_20" at 345,267 size 96x32; TextOff 'ON'
      Visibility <- "Motor_vibrador_tunel_1"
   Button "Button_21" at 469,268 size 96x32; TextOff 'OFF'
      Visibility <- "Motor_vibrador_tunel_1"
   Button "Button_22" at 604,268 size 96x32; TextOff 'FALLA'
      Visibility <- "Señal_de_fallo_vibrador_tunel_1"
   Button "Button_24" at 345,308 size 96x32; TextOff 'ABIERTA'
      Visibility <- "Subir_Cuchara_Tunel_1"
   Button "Button_25" at 469,309 size 96x32; TextOff 'CERRADA'
      Visibility <- "Bajar_cuchara_Tunel_1"
   Button "Button_28" at 345,352 size 96x32; TextOff 'DERECHA'
      Visibility <- "Desviar_cajas_derecha_Tunel_1"
   Button "Button_29" at 469,353 size 96x32; TextOff 'IZQUIERDA'
      Visibility <- "Desviar_cajas_izquierda_Tunel_1"
   GraphicView "Graphic view_2" at 729,118 size 35x35; Picture "ADVERTENCIA"
      Visibility <- "Señal_de_fallo_banda_tunel_1"
   GraphicView "Graphic view_3" at 729,166 size 35x35; Picture "ADVERTENCIA"
      Visibility <- "Señal_de_fallo_aspirador_tunel_1"
   GraphicView "Graphic view_4" at 729,214 size 35x35; Picture "ADVERTENCIA"
      Visibility <- "Señal_de_fallo_ventilador_tunel_1"
   GraphicView "Graphic view_5" at 729,264 size 35x35; Picture "ADVERTENCIA"
      Visibility <- "Señal_de_fallo_vibrador_tunel_1"
   GraphicView "Graphic view_1" at 0,0 size 100x100; Picture "pngegg"
   Button "Button_11" at 119,435 size 368x32; TextOff 'VISUALIZACION MIMICO'
      on Press: ActivateScreen("MODO REMOTO", 0)
   Button "Button_10" at 530,435 size 172x32; TextOff 'CONFIGURACION'; Authorization "Mantenimiento"
      on Press: ActivateScreen("VISUALIZACION DE ESTADOS LOCAL TUNEL 1", 0)
   UserView "User view_1" at 118,10 size 564x55
   Softkey "Softkey_F1" at 0,0 size 0x0
      on KeyDown: ActivateScreen("PANTALLA DE INICIO", 0)

screen "CONFIGURACION TUNEL 1" 800x480
   GraphicView "Graphic view_1" at 0,0 size 100x100; Picture "pngegg"
   GraphicView "Graphic view_29" at 712,14 size 60x60; Picture "Graphic_28"
      Visibility <- "Señalizacion_operacion_verde_tunel_1"
   GraphicView "Graphic view_30" at 714,14 size 60x60; Picture "Graphic_29"
      Visibility <- "Señalizacion_azul_tunel_1"
   GraphicView "Graphic view_31" at 716,14 size 60x60; Picture "Graphic_31"
      Visibility <- "Señalizacion_Roja_Tunel_1"
   IOField "I/O field_1" at 468,193 size 100x32; Authorization "Admon"; FormatPattern s999; Unit  Seg
      on Activate: function_bbf3fe93(1, N)
      ProcessValue <- "TEMPORIZADOR_PASO_TAPAS_TUNEL_1"
   IOField "I/O field_2" at 468,247 size 100x32; Authorization "Admon"; FormatPattern s999; Unit  Seg
      ProcessValue <- "TEMPORIZADOR_BLOQUEO_TAPAS_TUNEL_1"
   IOField "I/O field_3" at 468,301 size 100x32; Authorization "Admon"; FormatPattern s999; Unit  Seg
      ProcessValue <- "TEMPORIZADOR_CAMBIO_DE_LLENADO_CAJA_TUNEL_1"
   Button "Button_1" at 193,193 size 252x32; TextOff 'TIEMPO DE PASO TAPAS'
   Button "Button_2" at 193,247 size 252x32; TextOff 'TIEMPO DE BLOQUEO TAPAS'
   Button "Button_3" at 193,302 size 252x32; TextOff 'TIEMPO DE CAMBIO CAJA'
   Button "Button_11" at 400,440 size 368x32; TextOff 'ESTADO DE ELEMENTOS Y ACTUADORES'
      on Press: ActivateScreen("VISUALIZACION DE ESTADOS LOCAL TUNEL 1", 0)
   Button "Button_4" at 23,440 size 368x32; TextOff 'VISUALIZACION MIMICO'
      on Press: ActivateScreen("MODO REMOTO", 0)
   UserView "User view_1" at 118,10 size 564x55
   Softkey "Softkey_F1" at 0,0 size 0x0
      on KeyDown: ActivateScreen("PANTALLA DE INICIO", 0)

screen "ALARMAS" 800x480
   GraphicView "Graphic view_1" at 0,0 size 100x100; Picture "pngegg"
   GraphicView "Graphic view_29" at 712,14 size 60x60; Picture "Graphic_28"
      Visibility <- "Señalizacion_operacion_verde_tunel_1"
   GraphicView "Graphic view_30" at 714,14 size 60x60; Picture "Graphic_29"
      Visibility <- "Señalizacion_azul_tunel_1"
   GraphicView "Graphic view_31" at 716,14 size 60x60; Picture "Graphic_31"
      Visibility <- "Señalizacion_Roja_Tunel_1"
   UserView "User view_1" at 118,10 size 564x55
   AlarmView "Alarm view_1" at 0,98 size 799x378
*)

(* ===== HMI "HMI_RT_3" =====
system functions are stored by id; their names below are inferred from use

HMI tags "Default tag table"
   "Tag_ScreenNumber" : UInt, internal

Template "Template_1" 800x480
   Button "Exit" at 714,429 size 71x50; TextOff 'Exit'; PictureOff "ExitRuntime_KTP700_Basic_PN_TR"; PictureOn "ExitRuntime_KTP700_Basic_PN_TR"
      on Release: StopRuntime(0)
   Button "Log on" at 614,429 size 71x50; TextOff 'Log on'; PictureOff "Login_KTP700_Basic_PN_TR"; PictureOn "Login_KTP700_Basic_PN_TR"
      on Release: function_a2a04561()
   Button "Template_Button" at 514,429 size 71x50; TextOff 'Text'
   Button "Template_Button_1" at 414,429 size 71x50; TextOff 'Text'
   Button "Template_Button_2" at 314,429 size 71x50; TextOff 'Text'
   Button "Template_Button_3" at 214,429 size 71x50; TextOff 'Text'
   Button "Alarms" at 114,429 size 71x50; TextOff 'Alarms'; PictureOff "AlarmDisplay_KTP700_Basic_PN_TR"; PictureOn "AlarmDisplay_KTP700_Basic_PN_TR"
      on Release: function_ef3f5d25("Alarm window_Unacknowledged", -1)
   Button "Start screen" at 14,429 size 71x50; TextOff 'Start screen'; PictureOff "NavigateHome_KTP700_Basic_PN_TR"; PictureOn "NavigateHome_KTP700_Basic_PN_TR"
      on Release: ActivateScreen("Root screen", 0)
   SymbolicIOField "Symbolic_IO_Field_Screen" at 93,9 size 600x33; TextOff '0'; TextOn '1'; TextList "TextList_ScreenNames"
      ProcessValue <- "Tag_ScreenNumber"
      on Change: ActivateScreenByNumber("Tag_ScreenNumber", 0)
   DateTimeField "HmiScreenItemData" at 695,25 size 105x25
   DateTimeField "HmiScreenItemData_1" at 695,0 size 105x25
   GraphicView "Logo" at 0,0 size 91x51; Picture "Logo of HMI_1"

screen "Root screen" 800x480, template "Template_1"
   on GenerateScreen: SetTag("Tag_ScreenNumber", 1)
   TextField "HmiScreenItemData" at 80,225 size 640x25; Text 'Welcome to HMI_1 (KTP700 Basic+ PN)!'
*)